
           IF #stringBox[#i] = #lineBreak THEN
               #lineBox[#pLineBox] := "Trim"(#lineBox[#pLineBox]);
               #pLineBox := #pLineBox + 1;
               #lineBox[#pLineBox] := #lineBreak;
               #pLineBox := #pLineBox + 1;
           END_IF;


           IF #stringBox[#i] <> #lineBreak THEN

               IF #i = 0 THEN
                   #lengthTest := #stringBox[#i];
               END_IF;

               IF #i >= 1 THEN
                   #lengthTest := CONCAT_WSTRING(IN1 := #lineBox[#pLineBox],
                                                 IN2 := #space,
                                                 IN3 := #stringBox[#i]);
               END_IF;

               IF LEN(#lengthTest) <= #maxLength THEN
                   #lineBox[#pLineBox] := #lengthTest;
               END_IF;

               IF LEN(#lengthTest) > #maxLength THEN
                   #lineBox[#pLineBox] := "Trim"(#lineBox[#pLineBox]);
                   #lineBox[#pLineBox] := "Trim"(#lineBox[#pLineBox]);
                   #pLineBox := #pLineBox + 1;
                   #lineBox[#pLineBox] := #stringBox[#i];
               END_IF;
           END_IF;

       END_FOR;

       FOR #i := 0 TO 10 DO

           IF #lineBox[#i] = #space OR #lineBox[#i] = WString#'' THEN
               EXIT;
           END_IF;
           IF #i = 0 THEN
               #output := #lineBox[#i];
           END_IF;
           IF #i >= 1 THEN
               IF #lineBox[#i] = #lineBreak THEN
                   #output := #output;
               END_IF;
               IF #lineBox[#i] <> #lineBreak THEN
                   #output := CONCAT_WSTRING(IN1 := #output,
                                             IN2 := #lineBreak,
                                             IN3 := #lineBox[#i]);
               END_IF;
           END_IF;

       END_FOR;

       #output := "Trim"(#output);

   END_IF;

   #"Word Wrap" := #output;
END_FUNCTION

FUNCTION "Trim" : WString   // FC29, SCL
{ S7_Optimized_Access := 'TRUE' }
VERSION : 0.1
   VAR_INPUT
      wString : WString;
   END_VAR
   VAR_TEMP
      ret : WString;
   END_VAR
   VAR CONSTANT
      space : WString := WSTRING#' ';
   END_VAR
BEGIN
   #ret := #wString;
   IF LEFT(IN := #ret, L := 1) = #space THEN
       #ret := RIGHT(IN := #ret, L := LEN(#ret) - 1);
   END_IF;
   IF RIGHT(IN := #ret, L := 1) = #space THEN
       #ret := LEFT(IN := #ret, L := LEN(#ret) - 1);
   END_IF;
   #Trim := #ret;
END_FUNCTION

FUNCTION "Upper" : Void   // FC49, SCL
{ S7_Optimized_Access := 'TRUE' }
VERSION : 0.1
   VAR_IN_OUT
      "string" : Variant;
   END_VAR
   VAR_TEMP
      "type" : Bool;
      stringBox : String;
      status : Int;
      wStringBox : WString;
      charArr : Array[0..255] of Char;
      cntChar : UInt;
      pChar : Int;
   END_VAR
   VAR CONSTANT
      asciiLow : Char := 'a';
      asciiHigh : Char := 'z';
      asciiCaseOffset : Int := 32;
   END_VAR
BEGIN
   IF TypeOf(#string) = String THEN
       #status := MOVE_BLK_VARIANT(SRC := #string,
                                   COUNT := 1,
                                   SRC_INDEX := 0,
                                   DEST_INDEX := 0,
                                   DEST => #stringBox);
   ELSIF TypeOf(#string) = WString THEN
       #status := MOVE_BLK_VARIANT(SRC := #string,
                                   COUNT := 1,
                                   SRC_INDEX := 0,
                                   DEST_INDEX := 0,
                                   DEST => #wStringBox);
       #stringBox := WSTRING_TO_STRING(#wStringBox);
   ELSE
       RETURN;
   END_IF;

   Strg_TO_Chars(Strg := #stringBox,
                 pChars := 0,
                 Cnt => #cntChar,
                 Chars := #charArr);

   FOR #pChar := 0 TO UINT_TO_INT(#cntChar) - 1 DO
       IF #asciiLow <= #charArr[#pChar] AND #charArr[#pChar] <= #asciiHigh THEN
           #charArr[#pChar] := INT_TO_CHAR(CHAR_TO_INT(#charArr[#pChar]) - #asciiCaseOffset);
       END_IF;
   END_FOR;

   Chars_TO_Strg(Chars := #charArr,
                 pChars := 0,
                 Cnt := #cntChar,
                 Strg => #stringBox);

   IF TypeOf(#string) = String THEN
       #status := MOVE_BLK_VARIANT(SRC := #stringBox,
                                   COUNT := 1,
                                   SRC_INDEX := 0,
                                   DEST_INDEX := 0,
                                   DEST => #string);
   ELSIF TypeOf(#string) = WString THEN
       #wStringBox := STRING_TO_WSTRING(#stringBox);
       #status := MOVE_BLK_VARIANT(SRC := #wStringBox,
                                   COUNT := 1,
                                   SRC_INDEX := 0,
                                   DEST_INDEX := 0,
                                   DEST => #string);
   END_IF;
END_FUNCTION

// folder: Utilities/Table Navigation

FUNCTION_BLOCK "Table Nav"   // FB43, SCL
{ S7_Optimized_Access := 'TRUE' }
VERSION : 0.1
   VAR_INPUT
      tblData : Variant;
      tblDisp : Variant;
      tableNav : "Table Nav: HMI";
   END_VAR
   VAR_IN_OUT
      rowIndices : Variant;
   END_VAR
   VAR
      "inst Pulses: Table Nav" : "Table Nav: Pulses";
      r1 : DInt;
   END_VAR
   VAR_TEMP
      len : Struct
         tblData : DInt;
         tblDisp : DInt;
      END_STRUCT;
      offset : DInt;
      pulses : "Table Nav: PLC";
      RET_VAL : Int;
      retRowIndices : Array[0..#lenRetArr] of DInt;
   END_VAR
   VAR CONSTANT
      lenRetArr : DInt := 999;
   END_VAR
BEGIN
   REGION "DESCRIPTION"
       (*
       The function returns row indicies indicating the visible rows of a larger
       table determined by standard table navigation buttons.
       The function uses the variant data type to handle tables of any size.
       Rollover and rollunder features are built in.
       *)    
   END_REGION

   REGION "GET PRESS PULSES"    
       #"inst Pulses: Table Nav"(press := #tableNav,
                                 pulses=> #pulses);
   END_REGION

   REGION "RUN ON BUTTON PRESS"
       IF "Table Nav: Run Trigger"(#pulses) THEN

           REGION "GET ARRAY PARAMETERS"
               #len.tblData := UDINT_TO_DINT(CountOfElements(#tblData));
               #len.tblDisp := UDINT_TO_DINT(CountOfElements(#tblDisp));
           END_REGION

           REGION "CALCULATE OFFSET"
               #offset := "Table Nav: Calculate Offset"(pulses := #pulses,
                                                        lenTblData := #len.tblData,
                                                        lenTblDisp := #len.tblDisp,
                                                        r1 := #r1);
           END_REGION

           REGION "CALCULATE FIRST ROW"
               #r1 := "Table Nav: Get First Row"(lenTblData := #len.tblData,
                                                 offset := #offset,
                                                 r1 := #r1);
           END_REGION

           REGION "CALCUALTE ROW INDICIES"
               "Table Nav: Calc Row Indices"(lenTblData := #len.tblData,
                                             lenTblDisp := #len.tblDisp,
                                             r1 := #r1,
                                             rowIndicies := #retRowIndices);
           END_REGION

           REGION "RETURN ROW INDICIES"
               #RET_VAL := MOVE_BLK_VARIANT(SRC := #retRowIndices,
                                            COUNT := DINT_TO_UDINT(#len.tblDisp),
                                            SRC_INDEX := 0,
                                            DEST_INDEX := 0,
                                            DEST => #rowIndices);
           END_REGION

       END_IF;
   END_REGION
END_FUNCTION_BLOCK

FUNCTION_BLOCK "Table Nav: Pulses"   // FB44, SCL
{ S7_Optimized_Access := 'TRUE' }
VERSION : 0.1
   VAR_INPUT
      press : "Table Nav: HMI";
   END_VAR
   VAR_OUTPUT
      pulses : "Table Nav: PLC";
   END_VAR
   VAR
      old : "Table Nav: PLC";
   END_VAR
BEGIN
   REGION "EVALUATION"
       #pulses.top := #press.top.actuate AND NOT #old.top;
       #pulses.pageUp := #press.pageUp.actuate AND NOT #old.pageUp;
       #pulses.lineUp := #press.lineUp.actuate AND NOT #old.lineUp;
       #pulses.lineDown := #press.lineDown.actuate AND NOT #old.lineDown;
       #pulses.pageDown := #press.pageDown.actuate AND NOT #old.pageDown;
       #pulses.bottom := #press.bottom.actuate AND NOT #old.bottom;
   END_REGION

   REGION "CHANGE DETECTION"
       #old.top := #press.top.actuate;
       #old.pageUp := #press.pageUp.actuate;
       #old.lineUp := #press.lineUp.actuate;
       #old.lineDown := #press.lineDown.actuate;
       #old.pageDown := #press.pageDown.actuate;
       #old.bottom := #press.bottom.actuate;
   END_REGION
END_FUNCTION_BLOCK

FUNCTION "Table Nav: Get First Row" : DInt   // FC44, SCL
{ S7_Optimized_Access := 'TRUE' }
VERSION : 0.1
   VAR_INPUT
      lenTblData : DInt;
      offset : DInt;
      r1 : DInt;
   END_VAR
   VAR_TEMP
      newR1 : DInt;
      trgRun : Bool;
   END_VAR
BEGIN
   REGION "DESCRIPTION"
       (*
       The new first row of the table is calculated from the offset. 
       Rollover and rollunder are resolved for the first row.
       *)
   END_REGION

   REGION "COPY TO INTERNAL"
       #newR1 := #r1 + #offset;
   END_REGION

   REGION "ROLLUNDER"
       IF #newR1 < 0 THEN
           #newR1 := #newR1 + #lenTblData;
       END_IF;
   END_REGION

   REGION "ROLLOVER"
       IF #newR1 > #lenTblData THEN
           #newR1 := #newR1 - #lenTblData;
       END_IF;
   END_REGION

   REGION "OUTPUT"
       #"Table Nav: Get First Row" := #newR1;
   END_REGION
END_FUNCTION

FUNCTION "Table Nav: Calculate Offset" : DInt   // FC45, SCL
{ S7_Optimized_Access := 'TRUE' }
VERSION : 0.1
   VAR_INPUT
      lenTblData : DInt;
      lenTblDisp : DInt;
      pulses : "Table Nav: PLC";
      r1 : DInt;
   END_VAR
   VAR_TEMP
      retOffset : DInt;
   END_VAR
   // Ret_Val : offset from table row 1 from button
BEGIN
   REGION "DESCRIPTION"
       (*
       The offset from the first row of the table is calculated based on the button pressed.
       *)
   END_REGION

   REGION "TOP"
       IF #pulses.top THEN
           #retOffset := -1 * #r1;
       END_IF;
   END_REGION

   REGION "PAGE UP"
       IF #pulses.pageUp THEN
           #retOffset := -1 * #lenTblDisp;
       END_IF;
   END_REGION

   REGION "LINE UP"
       IF #pulses.lineUp THEN
           #retOffset := -1;
       END_IF;
   END_REGION

   REGION "LINE DOWN"
       IF #pulses.lineDown THEN
           #retOffset := 1;
       END_IF;
   END_REGION

   REGION "PAGE DOWN"
       IF #pulses.pageDown THEN
           #retOffset := #lenTblDisp ;
       END_IF;
   END_REGION

   REGION "BOTTOM"
       IF #pulses.bottom THEN
           #retOffset := #lenTblData - #lenTblDisp - #r1;
       END_IF;
   END_REGION

   REGION "RETURN"
       #"Table Nav: Calculate Offset" := #retOffset;
   END_REGION
END_FUNCTION

FUNCTION "Table Nav: Calc Row Indices" : Void   // FC46, SCL
{ S7_Optimized_Access := 'TRUE' }
VERSION : 0.1
   VAR_INPUT
      lenTblData : DInt;
      lenTblDisp : DInt;
      r1 : DInt;
   END_VAR
   VAR_IN_OUT
      rowIndicies : Array[0..#lenRetArr] of DInt;
   END_VAR
   VAR_TEMP
      pOutArr : Int;
      calcRowIdx : DInt;
      retRowIndicies : Array[0..#lenRetArr] of DInt;
   END_VAR
   VAR CONSTANT
      lenRetArr : DInt := 999;
   END_VAR
BEGIN
   REGION "DESCRIPTION"
       (*
       An array of the row indicies that the table should display is returned.
       Rollover and rollunder are calculated index by index.
       *) 
   END_REGION

   REGION "INITIALIZE OUTPUT"
       FOR #pOutArr := 0 TO #lenRetArr DO
           #rowIndicies[#pOutArr] := 0;
       END_FOR;
   END_REGION

   REGION "CALCULATE INDICIES"
       FOR #pOutArr := 0 TO #lenTblDisp DO

           REGION "CALCULATE INDEX"
               #calcRowIdx := #r1 + #pOutArr;
           END_REGION

           REGION "ROLL UNDER"
               IF #calcRowIdx < 0 THEN
                   #calcRowIdx := #calcRowIdx + #lenTblDisp;
               END_IF;
           END_REGION

           REGION "ROLL OVER"
               IF #calcRowIdx >= #lenTblData THEN
                   #calcRowIdx := #calcRowIdx - #lenTblData;
               END_IF;
           END_REGION

           REGION "SAVE TO ARRAY"
               #retRowIndicies[#pOutArr] := #calcRowIdx;
           END_REGION

       END_FOR;
   END_REGION

   REGION "OUTPUT"
       #rowIndicies := #retRowIndicies;
   END_REGION
END_FUNCTION

FUNCTION "Table Nav: Run Trigger" : Bool   // FC47, SCL
{ S7_Optimized_Access := 'TRUE' }
VERSION : 0.1
   VAR_INPUT
      pulses : "Table Nav: PLC";
   END_VAR
BEGIN
       #"Table Nav: Run Trigger" :=
       #pulses.top OR
       #pulses.pageUp OR
       #pulses.lineUp OR
       #pulses.lineDown OR
       #pulses.pageDown OR
       #pulses.bottom;
END_FUNCTION

// folder: Utilities/Timer

FUNCTION "Timer: Time to WString" : WString   // FC36, SCL
{ S7_Optimized_Access := 'TRUE' }
VERSION : 0.1
   VAR_INPUT
      "Time" : Time;
   END_VAR
   VAR_TEMP
      "Time as DInt" : DInt;
      "Hours 10s Place" : DInt;
      "Hours 1s Place" : DInt;
      "Minutes 10s Place" : DInt;
      "Minutes 1s Place" : DInt;
      "Seconds 10s Place" : DInt;
      "Seconds 1s Place" : DInt;
      "Time Elements" : Array[0..4] of WString;
      Length : Int;
      "String Box" : WString;
      "DInt Box" : DInt;
   END_VAR
   VAR CONSTANT
      "Milliseconds per 10 Hours" : DInt := 36_000_000;
      "Milliseconds per Hour" : DInt := 3_600_000;
      "Milliseconds per 10 Minutes" : DInt := 600_000;
      "Milliseconds per Minute" : DInt := 60_000;
      "Milliseconds per 10 Seconds" : DInt := 10_000;
      "Milliseconds per Second" : DInt := 1_000;
   END_VAR
BEGIN
   REGION GET INPUT
       #"Time as DInt" := #Time;
   END_REGION

   REGION CONVERT TIME INTO INDIVIDUAL PLACE VALUES
       #"Minutes 10s Place" := #"Time as DInt" / #"Milliseconds per 10 Minutes";
       #"Minutes 1s Place" := (#"Time as DInt" / #"Milliseconds per Minute") MOD 10;
       #"Seconds 10s Place" := (#"Time as DInt" MOD #"Milliseconds per Minute") / #"Milliseconds per 10 Seconds";
       #"Seconds 1s Place" := (#"Time as DInt" / #"Milliseconds per Second") MOD 10;
   END_REGION

   REGION "ADD SIGN"
       #"Time Elements"[0] := wstring#'';
       IF #"Minutes 10s Place" < 0 OR
           #"Minutes 1s Place" < 0 OR
           #"Seconds 10s Place" < 0 OR
           #"Seconds 1s Place" < 0 THEN
            #"Time Elements"[0] := wstring#'-';
       END_IF;
   END_REGION

   REGION CONVERT PLACE VALUES INTO COMPONENT STRINGS
       // MINUTES
       #"DInt Box" := #"Minutes 10s Place" * 10 + #"Minutes 1s Place";
       #"String Box" := DINT_TO_WSTRING(IN := #"DInt Box");
       #"String Box" := "Strip Sign"("WString":=#"String Box");
       #"String Box" := "Add Leading"("Leading Character" := WCHAR#'0',
                                      "Desired Length" := 2,
                                      "String" := #"String Box");
       #"Time Elements"[1] := #"String Box";
       // COLON
       #"Time Elements"[2] := WSTRING#':';
       // SECONDS
       #"DInt Box" := #"Seconds 10s Place" * 10 + #"Seconds 1s Place";
       #"String Box" := DINT_TO_WSTRING(IN := #"DInt Box");
       #"String Box" := "Strip Sign"("WString":=#"String Box");
       #"String Box" := "Add Leading"("Leading Character" := WCHAR#'0',
                                      "Desired Length" := 2,
                                      "String" := #"String Box");
       #"Time Elements"[3] := #"String Box";
   END_REGION


   REGION RETURN VALUE
       #"Timer: Time to WString" := CONCAT_WSTRING(IN1 := #"Time Elements"[0],
                                            IN2 := #"Time Elements"[1],
                                            IN3 := #"Time Elements"[2],
                                            IN4 := #"Time Elements"[3]);
   END_REGION
END_FUNCTION

FUNCTION "Timer: WString to Time" : Time   // FC38, SCL
{ S7_Optimized_Access := 'TRUE' }
VERSION : 0.1
   VAR_INPUT
      WString : WString;
   END_VAR
   VAR_TEMP
      Count : UInt;
      "DInt Box" : DInt;
      "String Box" : WString [5];
      "Time Box" : Time;
      "WChar Array" : Array[0..4] of WChar;
   END_VAR
   VAR CONSTANT
      "ms/(10 hr)" : DInt := 36_000_000;
      "ms/hr" : DInt := 3_600_000;
      "ms/(10 min)" : DInt := 600_000;
      "ms/min" : DInt := 60_000;
      "ms/(10 sec)" : DInt := 10_000;
      "ms/sec" : DInt := 1_000;
   END_VAR
BEGIN
   REGION EXPLODE INPUT

       #"String Box" := #WString;
       IF #"String Box" = WSTRING#'' THEN
           #"String Box" := WSTRING#'00:00';
       END_IF;

       Strg_TO_Chars(Strg := #"String Box",
                     pChars := 0,
                     Cnt => #Count,
                     Chars := #"WChar Array");

   END_REGION

   REGION CONVERT ARRAY ELEMENTS TO TIME

       // 10S OF MINUTES
       #"DInt Box" := WCHAR_TO_DINT(IN := #"WChar Array"[0]) - 16#30;
       #"Time Box" := #"Time Box" + #"DInt Box" * #"ms/(10 min)";

       // MINUTES
       #"DInt Box" := WCHAR_TO_DINT(IN := #"WChar Array"[1]) - 16#30;
       #"Time Box" := #"Time Box" + #"DInt Box" * #"ms/min";

       // 10S OF SECONDS
       #"DInt Box" := WCHAR_TO_DINT(IN := #"WChar Array"[3]) - 16#30;
       #"Time Box" := #"Time Box" + #"DInt Box" * #"ms/(10 sec)";

       // SECONDS
       #"DInt Box" := WCHAR_TO_DINT(IN := #"WChar Array"[4]) - 16#30;
       #"Time Box" := #"Time Box" + #"DInt Box" * #"ms/sec";

   END_REGION


   REGION RETURN VALUE

       #"Timer: WString to Time" := #"Time Box";

   END_REGION
END_FUNCTION

FUNCTION "Timer: WString to Real" : Real   // FC39, SCL
{ S7_Optimized_Access := 'TRUE' }
VERSION : 0.1
   VAR_INPUT
      wstring : WString;
   END_VAR
   VAR CONSTANT
      msPerSec : Real := 1000.0;
   END_VAR
BEGIN
   #"Timer: WString to Real" := DINT_TO_REAL(TIME_TO_DINT("Timer: WString to Time"(#wstring))) / #msPerSec;
END_FUNCTION

FUNCTION "Timer: Real to WString" : WString   // FC40, SCL
{ S7_Optimized_Access := 'TRUE' }
VERSION : 0.1
   VAR_INPUT
      realVal : Real;
   END_VAR
   VAR CONSTANT
      msPerSec : Real := 1000.0;
   END_VAR
BEGIN
   #"Timer: Real to WString" := "Timer: Time to WString"(DINT_TO_TIME(REAL_TO_DINT(#realVal * #msPerSec)));
END_FUNCTION

// ===== library types =====

TYPE "Table Row Data"
   STRUCT
      address : UInt;
      ordered : Bool;
      pbSelection : Struct
         actuate : Bool;
         animate : USInt;
      END_STRUCT;
      rtBackground : Struct
         animate : USInt;
      END_STRUCT;
      tfDropZone : Struct
         animate : USInt;
         value : WString[20];
      END_STRUCT;
      tfLine : Struct
         animate : USInt;
         value : WString[20];
      END_STRUCT;
      tfPartNumber : Struct
         animateDL : USInt;
         animateSL : USInt;
         value : WString[40];
      END_STRUCT;
      tfTime : Struct
         animate : USInt;
         value : WString[20];
      END_STRUCT;
   END_STRUCT;
END_TYPE

TYPE "Station Assignment: Button Details Data"
   STRUCT
      alloted : Struct
         animate : USInt;
         value : WString[10];
      END_STRUCT;
      critical : Struct
         animate : USInt;
         value : WString[10];
      END_STRUCT;
      label : Struct
         animate : USInt;
         value : WString[2];
      END_STRUCT;
      partNumber : Struct
         animate : USInt;
         value : WString[40];
      END_STRUCT;
      select : Struct
         actuate : Bool;
         animate : USInt;
      END_STRUCT;
   END_STRUCT;
END_TYPE

TYPE "Station Sim Data"
   STRUCT
      stn : Struct
         animate : USInt;
         label : WString[20];
      END_STRUCT;
      btn : Struct
         actuate : Byte;
         animate : Array[0..7] of USInt;
         labels : Array[0..7] of WString [4];
      END_STRUCT;
   END_STRUCT;
END_TYPE

(* ===== HMI "HMI_RT_1" =====
system functions are stored by id; their names below are inferred from use
connection "Main HMI": ETHERNET, S7_1500_OMS

HMI tags "Default tag table"
   "Clock_Byte" : Byte = PLC Clock_Byte AT %MB0, 100 ms
   "HMI_screenNumber" : Int = PLC HMI.screenNumber AT %DB1.DBW0, 100 ms
   "HMI_barcode" : Barcode Screen = PLC HMI.barcode AT %DB1.DBW0, 100 ms
   "HMI_partCall_row{0}" : Table Row = PLC HMI.partCall.row[0], 100 ms
   "HMI_partCall_row{1}" : Table Row = PLC HMI.partCall.row[1], 100 ms
   "HMI_partCall_row{2}" : Table Row = PLC HMI.partCall.row[2], 100 ms
   "HMI_partCall_row{3}" : Table Row = PLC HMI.partCall.row[3], 100 ms
   "HMI_partCall_row{4}" : Table Row = PLC HMI.partCall.row[4], 100 ms
   "HMI_partCall_row{5}" : Table Row = PLC HMI.partCall.row[5], 100 ms
   "HMI_partCall_row{6}" : Table Row = PLC HMI.partCall.row[6], 100 ms
   "HMI_partCall_row{7}" : Table Row = PLC HMI.partCall.row[7], 100 ms
   "HMI_partCall_row{8}" : Table Row = PLC HMI.partCall.row[8], 100 ms
   "HMI_partCall_row{9}" : Table Row = PLC HMI.partCall.row[9], 100 ms
   "HMI_partCall_row{10}" : Table Row = PLC HMI.partCall.row[10], 100 ms
   "HMI_settings_stations_selectBtns{0}" : PB Data: Text Label = PLC HMI.settings.stations.selectBtns[0], 100 ms
   "HMI_settings_stations_selectBtns{1}" : PB Data: Text Label = PLC HMI.settings.stations.selectBtns[1], 100 ms
   "HMI_settings_stations_selectBtns{2}" : PB Data: Text Label = PLC HMI.settings.stations.selectBtns[2], 100 ms
   "HMI_settings_stations_selectBtns{3}" : PB Data: Text Label = PLC HMI.settings.stations.selectBtns[3], 100 ms
   "HMI_settings_stations_selectBtns{4}" : PB Data: Text Label = PLC HMI.settings.stations.selectBtns[4], 100 ms
   "HMI_settings_stations_selectBtns{5}" : PB Data: Text Label = PLC HMI.settings.stations.selectBtns[5], 100 ms
   "HMI_settings_stations_selectBtns{6}" : PB Data: Text Label = PLC HMI.settings.stations.selectBtns[6], 100 ms
   "HMI_settings_stations_selectBtns{7}" : PB Data: Text Label = PLC HMI.settings.stations.selectBtns[7], 100 ms
   "HMI_settings_stations_selectBtns{8}" : PB Data: Text Label = PLC HMI.settings.stations.selectBtns[8], 100 ms
   "HMI_settings_stations_selectBtns{9}" : PB Data: Text Label = PLC HMI.settings.stations.selectBtns[9], 100 ms
   "HMI_settings_stations_selectBtns{10}" : PB Data: Text Label = PLC HMI.settings.stations.selectBtns[10], 100 ms
   "HMI_settings_stations_selectBtns{11}" : PB Data: Text Label = PLC HMI.settings.stations.selectBtns[11], 100 ms
   "HMI_settings_kp8_buttons{0}" : PB Data: Text Label = PLC HMI.settings.kp8.buttons[0], 100 ms
   "HMI_settings_kp8_buttons{7}" : PB Data: Text Label = PLC HMI.settings.kp8.buttons[7], 100 ms
   "HMI_settings_kp8_buttons{3}" : PB Data: Text Label = PLC HMI.settings.kp8.buttons[3], 100 ms
   "HMI_settings_kp8_buttons{6}" : PB Data: Text Label = PLC HMI.settings.kp8.buttons[6], 100 ms
   "HMI_settings_kp8_buttons{2}" : PB Data: Text Label = PLC HMI.settings.kp8.buttons[2], 100 ms
   "HMI_settings_kp8_buttons{5}" : PB Data: Text Label = PLC HMI.settings.kp8.buttons[5], 100 ms
   "HMI_settings_kp8_buttons{1}" : PB Data: Text Label = PLC HMI.settings.kp8.buttons[1], 100 ms
   "HMI_settings_kp8_buttons{4}" : PB Data: Text Label = PLC HMI.settings.kp8.buttons[4], 100 ms
   "HMI_settings_stations_selCount" : Int = PLC HMI.settings.stations.selCount, 100 ms
   "HMI_settings_viewingStation_btns{0}" : Station: Assignment: Button Details = PLC HMI.settings.viewingStation.btns[0], 100 ms
   "HMI_settings_viewingStation_btns{1}" : Station: Assignment: Button Details = PLC HMI.settings.viewingStation.btns[1], 100 ms
   "HMI_settings_viewingStation_btns{2}" : Station: Assignment: Button Details = PLC HMI.settings.viewingStation.btns[2], 100 ms
   "HMI_settings_viewingStation_btns{3}" : Station: Assignment: Button Details = PLC HMI.settings.viewingStation.btns[3], 100 ms
   "HMI_settings_viewingStation_btns{4}" : Station: Assignment: Button Details = PLC HMI.settings.viewingStation.btns[4], 100 ms
   "HMI_settings_viewingStation_btns{5}" : Station: Assignment: Button Details = PLC HMI.settings.viewingStation.btns[5], 100 ms
   "HMI_settings_viewingStation_previous" : PB Data: Graphic/Text List = PLC HMI.settings.viewingStation.previous, 100 ms
   "HMI_settings_viewingStation_next" : PB Data: Graphic/Text List = PLC HMI.settings.viewingStation.next, 100 ms
   "HMI_settings_stations_selectAll" : PB Data: Text Label = PLC HMI.settings.stations.selectAll, 100 ms
   "HMI_settings_partNumber_assign" : PB Data: Text Label = PLC HMI.settings.partNumber.assign, 100 ms
   "HMI_settings_partNumber_ioField" : IO Field Data: Part Number = PLC HMI.settings.partNumber.ioField, 100 ms
   "HMI_settings_alotted_assign" : PB Data: Text Label = PLC HMI.settings.alotted.assign, 100 ms
   "HMI_settings_alotted_ioField" : IO Field Data: Timers = PLC HMI.settings.alotted.ioField, 100 ms
   "HMI_settings_critical_assign" : PB Data: Text Label = PLC HMI.settings.critical.assign, 100 ms
   "HMI_settings_critical_ioField" : IO Field Data: Timers = PLC HMI.settings.critical.ioField, 100 ms
   "HMI_settings_kp8_selectButtons" : PB Data: Text Label = PLC HMI.settings.kp8.selectButtons, 100 ms
   "HMI_settings_viewingStation_dzData" : Drop Zone Data = PLC HMI.settings.viewingStation.dzData, 100 ms
   "HMI_settings_viewingStation_lineData" : Line Label Data = PLC HMI.settings.viewingStation.lineData, 100 ms
   "HMI_settings_stations_prevGroup" : PB Data: Graphic/Text List = PLC HMI.settings.stations.prevGroup, 100 ms
   "HMI_settings_stations_nextGroup" : PB Data: Graphic/Text List = PLC HMI.settings.stations.nextGroup, 100 ms
   "HMI_settings_viewingStation_name" : WString[20] = PLC HMI.settings.viewingStation.name, 100 ms
   "HMI_tableNav_top" : PB Data: Graphic/Text List = PLC HMI.tableNav.top, 100 ms
   "HMI_tableNav_pageUp" : PB Data: Graphic/Text List = PLC HMI.tableNav.pageUp, 100 ms
   "HMI_tableNav_lineUp" : PB Data: Graphic/Text List = PLC HMI.tableNav.lineUp, 100 ms
   "HMI_tableNav_lineDown" : PB Data: Graphic/Text List = PLC HMI.tableNav.lineDown, 100 ms
   "HMI_tableNav_pageDown" : PB Data: Graphic/Text List = PLC HMI.tableNav.pageDown, 100 ms
   "HMI_tableNav_bottom" : PB Data: Graphic/Text List = PLC HMI.tableNav.bottom, 100 ms
   "HMI_simStations_stations{0}" : Station: Sim Data = PLC HMI.simStations.me[0] AT %DB1.DBX0.0, 100 ms
   "HMI_simStations_me{1}" : Station: Sim Data = PLC HMI.simStations.me[1], 100 ms
   "HMI_simStations_me{2}" : Station: Sim Data = PLC HMI.simStations.me[2], 100 ms
   "HMI_simStations_me{3}" : Station: Sim Data = PLC HMI.simStations.me[3], 100 ms
   "HMI_simStations_me{4}" : Station: Sim Data = PLC HMI.simStations.me[4], 100 ms
   "HMI_simStations_me{5}" : Station: Sim Data = PLC HMI.simStations.me[5], 100 ms
   "HMI_simStations_me{6}" : Station: Sim Data = PLC HMI.simStations.me[6], 100 ms
   "HMI_simStations_me{7}" : Station: Sim Data = PLC HMI.simStations.me[7], 100 ms
   "HMI_simStations_me{8}" : Station: Sim Data = PLC HMI.simStations.me[8], 100 ms
   "HMI_simStations_me{9}" : Station: Sim Data = PLC HMI.simStations.me[9], 100 ms
   "HMI_simStations_me{10}" : Station: Sim Data = PLC HMI.simStations.me[10], 100 ms
   "HMI_simStations_me{11}" : Station: Sim Data = PLC HMI.simStations.me[11], 100 ms
   "HMI_simStations_up" : PB Data: Graphic/Text List = PLC HMI.simStations.up, 100 ms
   "HMI_simStations_down" : PB Data: Graphic/Text List = PLC HMI.simStations.down, 100 ms
   "HMI_networkHealth_pnioDevices{1}" : PB Data: Text Label = PLC HMI.networkHealth.pnioDevices[1], 100 ms
   "HMI_networkHealth_pnioDevices{2}" : PB Data: Text Label = PLC HMI.networkHealth.pnioDevices[2], 100 ms
   "HMI_networkHealth_pnioDevices{3}" : PB Data: Text Label = PLC HMI.networkHealth.pnioDevices[3], 100 ms
   "HMI_networkHealth_pnioDevices{4}" : PB Data: Text Label = PLC HMI.networkHealth.pnioDevices[4], 100 ms
   "HMI_networkHealth_pnioDevices{5}" : PB Data: Text Label = PLC HMI.networkHealth.pnioDevices[5], 100 ms
   "HMI_networkHealth_pnioDevices{6}" : PB Data: Text Label = PLC HMI.networkHealth.pnioDevices[6], 100 ms
   "HMI_networkHealth_pnioDevices{7}" : PB Data: Text Label = PLC HMI.networkHealth.pnioDevices[7], 100 ms
   "HMI_networkHealth_pnioDevices{8}" : PB Data: Text Label = PLC HMI.networkHealth.pnioDevices[8], 100 ms
   "HMI_networkHealth_pnioDevices{9}" : PB Data: Text Label = PLC HMI.networkHealth.pnioDevices[9], 100 ms
   "HMI_networkHealth_pnioDevices{10}" : PB Data: Text Label = PLC HMI.networkHealth.pnioDevices[10], 100 ms
   "HMI_networkHealth_pnioDevices{11}" : PB Data: Text Label = PLC HMI.networkHealth.pnioDevices[11], 100 ms
   "HMI_networkHealth_pnioDevices{12}" : PB Data: Text Label = PLC HMI.networkHealth.pnioDevices[12], 100 ms
   "HMI_networkHealth_pnioDevices{13}" : PB Data: Text Label = PLC HMI.networkHealth.pnioDevices[13], 100 ms
   "HMI_networkHealth_pnioDevices{16}" : PB Data: Text Label = PLC HMI.networkHealth.pnioDevices[16], 100 ms
   "HMI_networkHealth_pnioDevices{14}" : PB Data: Text Label = PLC HMI.networkHealth.pnioDevices[14], 100 ms
   "HMI_networkHealth_pnioDevices{15}" : PB Data: Text Label = PLC HMI.networkHealth.pnioDevices[15], 100 ms
   "HMI_networkHealth_pnioDevices{17}" : PB Data: Text Label = PLC HMI.networkHealth.pnioDevices[17], 100 ms
   "HMI_networkHealth_pnioDevices{18}" : PB Data: Text Label = PLC HMI.networkHealth.pnioDevices[18], 100 ms
   "HMI_networkHealth_pnioDevices{19}" : PB Data: Text Label = PLC HMI.networkHealth.pnioDevices[19], 100 ms
   "HMI_networkHealth_pnioDevices{20}" : PB Data: Text Label = PLC HMI.networkHealth.pnioDevices[20], 100 ms
   "HMI_networkHealth_pnioDevices{21}" : PB Data: Text Label = PLC HMI.networkHealth.pnioDevices[21], 100 ms
   "HMI_networkHealth_pnioDevices{22}" : PB Data: Text Label = PLC HMI.networkHealth.pnioDevices[22], 100 ms
   "HMI_networkHealth_pnioDevices{31}" : PB Data: Text Label = PLC HMI.networkHealth.pnioDevices[31], 100 ms
   "HMI_networkHealth_pnioDevices{32}" : PB Data: Text Label = PLC HMI.networkHealth.pnioDevices[32], 100 ms
   "HMI_networkHealth_pnioDevices{29}" : PB Data: Text Label = PLC HMI.networkHealth.pnioDevices[29], 100 ms
   "HMI_networkHealth_pnioDevices{30}" : PB Data: Text Label = PLC HMI.networkHealth.pnioDevices[30], 100 ms
   "HMI_networkHealth_pnioDevices{27}" : PB Data: Text Label = PLC HMI.networkHealth.pnioDevices[27], 100 ms
   "HMI_networkHealth_pnioDevices{28}" : PB Data: Text Label = PLC HMI.networkHealth.pnioDevices[28], 100 ms
   "HMI_networkHealth_pnioDevices{23}" : PB Data: Text Label = PLC HMI.networkHealth.pnioDevices[23], 100 ms
   "HMI_networkHealth_pnioDevices{24}" : PB Data: Text Label = PLC HMI.networkHealth.pnioDevices[24], 100 ms
   "HMI_networkHealth_pnioDevices{25}" : PB Data: Text Label = PLC HMI.networkHealth.pnioDevices[25], 100 ms
   "HMI_networkHealth_pnioDevices{26}" : PB Data: Text Label = PLC HMI.networkHealth.pnioDevices[26], 100 ms
   "HMI_networkHealth_pnioDevices{33}" : PB Data: Text Label = PLC HMI.networkHealth.pnioDevices[33], 100 ms
   "HMI_networkHealth_pnioDevices{34}" : PB Data: Text Label = PLC HMI.networkHealth.pnioDevices[34], 100 ms
   "HMI_networkHealth_pnioDevices{35}" : PB Data: Text Label = PLC HMI.networkHealth.pnioDevices[35], 100 ms
   "HMI_networkHealth_pnioDevices{36}" : PB Data: Text Label = PLC HMI.networkHealth.pnioDevices[36], 100 ms
   "HMI_networkHealth_pnioDevices{37}" : PB Data: Text Label = PLC HMI.networkHealth.pnioDevices[37], 100 ms
   "HMI_networkHealth_pnioDevices{38}" : PB Data: Text Label = PLC HMI.networkHealth.pnioDevices[38], 100 ms
   "HMI_networkHealth_pnioDevices{39}" : PB Data: Text Label = PLC HMI.networkHealth.pnioDevices[39], 100 ms
   "HMI_networkHealth_pnioDevices{40}" : PB Data: Text Label = PLC HMI.networkHealth.pnioDevices[40], 100 ms
   "HMI_networkHealth_pnioDevices{41}" : PB Data: Text Label = PLC HMI.networkHealth.pnioDevices[41], 100 ms
   "HMI_networkHealth_pnioDevices{42}" : PB Data: Text Label = PLC HMI.networkHealth.pnioDevices[42], 100 ms
   "HMI_networkHealth_pnioDevices{43}" : PB Data: Text Label = PLC HMI.networkHealth.pnioDevices[43], 100 ms
   "HMI_networkHealth_pnioDevices{44}" : PB Data: Text Label = PLC HMI.networkHealth.pnioDevices[44], 100 ms
   "HMI_networkHealth_pnioDevices{45}" : PB Data: Text Label = PLC HMI.networkHealth.pnioDevices[45], 100 ms
   "HMI_networkHealth_pnioDevices{46}" : PB Data: Text Label = PLC HMI.networkHealth.pnioDevices[46], 100 ms
   "HMI_networkHealth_pnioDevices{47}" : PB Data: Text Label = PLC HMI.networkHealth.pnioDevices[47], 100 ms
   "HMI_networkHealth_pnioDevices{48}" : PB Data: Text Label = PLC HMI.networkHealth.pnioDevices[48], 100 ms
   "HMI_networkHealth_et200spPopUp" : Station: ET200SP Comm Debug Data = PLC HMI.networkHealth.et200spPopUp, 100 ms
   "HMI_networkHealth_kp8PopUp" : Station: KP8 Comm Debug Data = PLC HMI.networkHealth.kp8PopUp, 100 ms
   "HMI_networkHealth_selectedDevice" : Int = PLC HMI.networkHealth.selectedDevice, 100 ms
   "Recipe Buffer_dropZone" : USInt = PLC "Recipe Buffer".dropZone, 1 s
   "Recipe Buffer_kp8Output" : DWord = PLC "Recipe Buffer".kp8Output, 1 s
   "Recipe Buffer_kp8LogicalState0" : Bool = PLC "Recipe Buffer".kp8LogicalState0, 1 s
   "Recipe Buffer_kp8LogicalState1" : Bool = PLC "Recipe Buffer".kp8LogicalState1, 1 s
   "Recipe Buffer_kp8LogicalState2" : Bool = PLC "Recipe Buffer".kp8LogicalState2, 1 s
   "Recipe Buffer_kp8LogicalState3" : Bool = PLC "Recipe Buffer".kp8LogicalState3, 1 s
   "Recipe Buffer_kp8LogicalState4" : Bool = PLC "Recipe Buffer".kp8LogicalState4, 1 s
   "Recipe Buffer_kp8LogicalState5" : Bool = PLC "Recipe Buffer".kp8LogicalState5, 1 s
   "Recipe Buffer_kp8LogicalState6" : Bool = PLC "Recipe Buffer".kp8LogicalState6, 1 s
   "Recipe Buffer_kp8LogicalState7" : Bool = PLC "Recipe Buffer".kp8LogicalState7, 1 s
   "Recipe Buffer_lineName" : USInt = PLC "Recipe Buffer".lineName, 1 s
   "Recipe Buffer_pnCode" : DInt = PLC "Recipe Buffer".pnCode, 1 s
   "Recipe Buffer_stackLight" : DWord = PLC "Recipe Buffer".stackLight, 1 s
   "Recipe Buffer_wipName" : WString[254] = PLC "Recipe Buffer".wipName, 1 s
   "Recipe Buffer_wipNumber" : UInt = PLC "Recipe Buffer".wipNumber, 1 s

text list "Station Selection Single": 0 'Select a Station to View'; 1 'Assignments'

recipe "Station01": dz <- "Recipe Buffer_dropZone", kp8Output <- "Recipe Buffer_kp8Output", logicalState0 <- "Recipe Buffer_kp8LogicalState0", logicalState1 <- "Recipe Buffer_kp8LogicalState1", logicalState2 <- "Recipe Buffer_kp8LogicalState2", logicalState3 <- "Recipe Buffer_kp8LogicalState3", logicalState4 <- "Recipe Buffer_kp8LogicalState4", logicalState5 <- "Recipe Buffer_kp8LogicalState5", logicalState6 <- "Recipe Buffer_kp8LogicalState6", logicalState7 <- "Recipe Buffer_kp8LogicalState7", lineName <- "Recipe Buffer_lineName", pnCode <- "Recipe Buffer_pnCode", stackLight <- "Recipe Buffer_stackLight", wipName <- "Recipe Buffer_wipName", wipNumber <- "Recipe Buffer_wipNumber"

recipe "Station02": dz <- "Recipe Buffer_dropZone", kp8Output <- "Recipe Buffer_kp8Output", logicalState0 <- "Recipe Buffer_kp8LogicalState0", logicalState1 <- "Recipe Buffer_kp8LogicalState1", logicalState2 <- "Recipe Buffer_kp8LogicalState2", logicalState3 <- "Recipe Buffer_kp8LogicalState3", logicalState4 <- "Recipe Buffer_kp8LogicalState4", logicalState5 <- "Recipe Buffer_kp8LogicalState5", logicalState6 <- "Recipe Buffer_kp8LogicalState6", logicalState7 <- "Recipe Buffer_kp8LogicalState7", lineName <- "Recipe Buffer_lineName", pnCode <- "Recipe Buffer_pnCode", stackLight <- "Recipe Buffer_stackLight", wipName <- "Recipe Buffer_wipName", wipNumber <- "Recipe Buffer_wipNumber"

recipe "Station03": dz <- "Recipe Buffer_dropZone", kp8Output <- "Recipe Buffer_kp8Output", logicalState0 <- "Recipe Buffer_kp8LogicalState0", logicalState1 <- "Recipe Buffer_kp8LogicalState1", logicalState2 <- "Recipe Buffer_kp8LogicalState2", logicalState3 <- "Recipe Buffer_kp8LogicalState3", logicalState4 <- "Recipe Buffer_kp8LogicalState4", logicalState5 <- "Recipe Buffer_kp8LogicalState5", logicalState6 <- "Recipe Buffer_kp8LogicalState6", logicalState7 <- "Recipe Buffer_kp8LogicalState7", lineName <- "Recipe Buffer_lineName", pnCode <- "Recipe Buffer_pnCode", stackLight <- "Recipe Buffer_stackLight", wipName <- "Recipe Buffer_wipName", wipNumber <- "Recipe Buffer_wipNumber"

recipe "Station04": dz <- "Recipe Buffer_dropZone", kp8Output <- "Recipe Buffer_kp8Output", logicalState0 <- "Recipe Buffer_kp8LogicalState0", logicalState1 <- "Recipe Buffer_kp8LogicalState1", logicalState2 <- "Recipe Buffer_kp8LogicalState2", logicalState3 <- "Recipe Buffer_kp8LogicalState3", logicalState4 <- "Recipe Buffer_kp8LogicalState4", logicalState5 <- "Recipe Buffer_kp8LogicalState5", logicalState6 <- "Recipe Buffer_kp8LogicalState6", logicalState7 <- "Recipe Buffer_kp8LogicalState7", lineName <- "Recipe Buffer_lineName", pnCode <- "Recipe Buffer_pnCode", stackLight <- "Recipe Buffer_stackLight", wipName <- "Recipe Buffer_wipName", wipNumber <- "Recipe Buffer_wipNumber"

recipe "Station05": dz <- "Recipe Buffer_dropZone", kp8Output <- "Recipe Buffer_kp8Output", logicalState0 <- "Recipe Buffer_kp8LogicalState0", logicalState1 <- "Recipe Buffer_kp8LogicalState1", logicalState2 <- "Recipe Buffer_kp8LogicalState2", logicalState3 <- "Recipe Buffer_kp8LogicalState3", logicalState4 <- "Recipe Buffer_kp8LogicalState4", logicalState5 <- "Recipe Buffer_kp8LogicalState5", logicalState6 <- "Recipe Buffer_kp8LogicalState6", logicalState7 <- "Recipe Buffer_kp8LogicalState7", lineName <- "Recipe Buffer_lineName", pnCode <- "Recipe Buffer_pnCode", stackLight <- "Recipe Buffer_stackLight", wipName <- "Recipe Buffer_wipName", wipNumber <- "Recipe Buffer_wipNumber"

recipe "Station06": dz <- "Recipe Buffer_dropZone", kp8Output <- "Recipe Buffer_kp8Output", logicalState0 <- "Recipe Buffer_kp8LogicalState0", logicalState1 <- "Recipe Buffer_kp8LogicalState1", logicalState2 <- "Recipe Buffer_kp8LogicalState2", logicalState3 <- "Recipe Buffer_kp8LogicalState3", logicalState4 <- "Recipe Buffer_kp8LogicalState4", logicalState5 <- "Recipe Buffer_kp8LogicalState5", logicalState6 <- "Recipe Buffer_kp8LogicalState6", logicalState7 <- "Recipe Buffer_kp8LogicalState7", lineName <- "Recipe Buffer_lineName", pnCode <- "Recipe Buffer_pnCode", stackLight <- "Recipe Buffer_stackLight", wipName <- "Recipe Buffer_wipName", wipNumber <- "Recipe Buffer_wipNumber"

screen "1 PART CALL" 1366x768
   on GenerateScreen: SetTag("HMI_screenNumber", 1)
   Rectangle "Settings Tab Background" at 682,0 size 684x68
      Appearance <- "HMI_screenNumber"
   Rectangle "Part Call Tab Background" at 0,0 size 685x68
      Appearance <- "HMI_screenNumber"
   Rectangle "Settings Tab Border Hide" at 685,61 size 678x20
      Visibility <- "HMI_screenNumber"
   Rectangle "Part Call Tab Border Hide" at 3,61 size 679x20
      Visibility <- "HMI_screenNumber"
   Button "Settings Screen" at 683,0 size 683x68; TextOff 'SETTINGS'; Authorization "User administration"
      on Release: ActivateScreen("2 SETTINGS", 0)
   Button "Part Call Screen" at 0,0 size 683x68; TextOff 'PART CALL'
      on Release: ActivateScreen("1 PART CALL", 0)
   TextField "Header Line" at 32,112 size 216x53; Text 'LINE'
   TextField "Header Drop Zone" at 238,112 size 236x53; Text 'DROP ZONE'
   TextField "Header Part Number" at 474,112 size 648x53; Text 'PART NUMBER'
   TextField "Header Time" at 1112,112 size 222x53; Text 'TIME'
   ScreenModuleView "TableRow00" at 27,170 size 1312x52; ScreenModuleType ""
      Guid_{11997190-27688} <- "HMI_partCall_row{0}"
      on Guid_{11997190-83214}: ActivateScreen("3 BARCODE", 0)
   ScreenModuleView "TableRow01" at 27,222 size 1312x52; ScreenModuleType ""
      Guid_{11997190-27688} <- "HMI_partCall_row{1}"
      on Guid_{11997190-83214}: ActivateScreen("3 BARCODE", 0)
   ScreenModuleView "TableRow02" at 27,274 size 1312x52; ScreenModuleType ""
      Guid_{11997190-27688} <- "HMI_partCall_row{2}"
      on Guid_{11997190-83214}: ActivateScreen("3 BARCODE", 0)
   ScreenModuleView "TableRow03" at 27,326 size 1312x52; ScreenModuleType ""
      Guid_{11997190-27688} <- "HMI_partCall_row{3}"
      on Guid_{11997190-83214}: ActivateScreen("3 BARCODE", 0)
   ScreenModuleView "TableRow04" at 27,378 size 1312x52; ScreenModuleType ""
      Guid_{11997190-27688} <- "HMI_partCall_row{4}"
      on Guid_{11997190-83214}: ActivateScreen("3 BARCODE", 0)
   ScreenModuleView "TableRow05" at 27,430 size 1312x52; ScreenModuleType ""
      Guid_{11997190-27688} <- "HMI_partCall_row{5}"
      on Guid_{11997190-83214}: ActivateScreen("3 BARCODE", 0)
   ScreenModuleView "TableRow06" at 27,482 size 1312x52; ScreenModuleType ""
      Guid_{11997190-27688} <- "HMI_partCall_row{6}"
      on Guid_{11997190-83214}: ActivateScreen("3 BARCODE", 0)
   ScreenModuleView "TableRow07" at 27,534 size 1312x52; ScreenModuleType ""
      Guid_{11997190-27688} <- "HMI_partCall_row{7}"
      on Guid_{11997190-83214}: ActivateScreen("3 BARCODE", 0)
   ScreenModuleView "TableRow08" at 27,586 size 1312x52; ScreenModuleType ""
      Guid_{11997190-27688} <- "HMI_partCall_row{8}"
      on Guid_{11997190-83214}: ActivateScreen("3 BARCODE", 0)
   ScreenModuleView "TableRow09" at 27,638 size 1312x52; ScreenModuleType ""
      Guid_{11997190-27688} <- "HMI_partCall_row{9}"
      on Guid_{11997190-83214}: ActivateScreen("3 BARCODE", 0)
   ScreenModuleView "TableRow10" at 27,690 size 1312x52; ScreenModuleType ""
      Guid_{11997190-27688} <- "HMI_partCall_row{10}"
      on Guid_{11997190-83214}: ActivateScreen("3 BARCODE", 0)

screen "2 SETTINGS" 1366x768
   on GenerateScreen: SetTag("HMI_screenNumber", 2)
   Rectangle "Part Call Nave Panel" at 0,0 size 455x68
      Appearance <- "HMI_screenNumber"
   Rectangle "Settings Nav Panel" at 452,0 size 462x68
      Appearance <- "HMI_screenNumber"
   Rectangle "Network Health Nav Panel" at 911,0 size 455x68
      Appearance <- "HMI_screenNumber"
   Rectangle "Part Call Border Hide" at 3,60 size 449x20
      Visibility <- "HMI_screenNumber"
   Rectangle "Settings Border Hide" at 455,60 size 456x20
      Visibility <- "HMI_screenNumber"
   Rectangle "Network Health Border Hide" at 914,60 size 449x20
      Visibility <- "HMI_screenNumber"
   Button "Part Call Screen" at 0,0 size 455x68; TextOff 'PART CALL'
      on Release: ActivateScreen("1 PART CALL", 0)
   Button "Settings Screen" at 455,0 size 460x68; TextOff 'SETTINGS'
      on Release: ActivateScreen("2 SETTINGS", 0)
   Button "Network Health Screen" at 914,0 size 452x68; TextOff 'NW HEALTH'
      on Release: ActivateScreen("4 NETWORK HEALTH", 0)
   Rectangle "Station Assignment Table BG Full" at 793,120 size 533x630
      Visibility <- "HMI_settings_stations_selCount"
   TextField "Current Station Single" at 803,130 size 513x45; Text 'Text'
      Visibility <- "HMI_settings_stations_selCount"
   TextField "Hide Line and Drop Zone Multi" at 803,181 size 513x40; Text 'select single station for Line and Drop Zone'
      Visibility <- "HMI_settings_stations_selCount"
   GraphicView "KP8 Image" at 496,327 size 275x412; Picture "kp8 image"
   Rectangle "Station Assignment Table BG Mini" at 793,120 size 533x65
      Visibility <- "HMI_settings_stations_selCount"
   ScreenModuleView "PB: Set PN" at 50,130 size 414x45; Guid_{11997190-63616} 'Assign Part Number'; ScreenModuleType ""
      Guid_{11997190-63605} <- "HMI_settings_partNumber_assign"
   ScreenModuleView "PN IO Field" at 50,180 size 414x50; ScreenModuleType ""
      Guid_{11997190-63113} <- "HMI_settings_partNumber_ioField"
   ScreenModuleView "PB: Set Allotted" at 494,130 size 137x45; Guid_{11997190-63616} 'Allotted'; ScreenModuleType ""
      Guid_{11997190-63605} <- "HMI_settings_alotted_assign"
   ScreenModuleView "PB: Set Critical" at 636,130 size 137x45; Guid_{11997190-63616} 'Crititcal'; ScreenModuleType ""
      Guid_{11997190-63605} <- "HMI_settings_critical_assign"
   ScreenModuleView "Alotted Time IO Field" at 494,180 size 137x50; ScreenModuleType ""
      Guid_{11997190-63269} <- "HMI_settings_alotted_ioField"
   ScreenModuleView "Critical Time IO Field" at 636,180 size 137x50; ScreenModuleType ""
      Guid_{11997190-63269} <- "HMI_settings_critical_ioField"
   ScreenModuleView "PB: Select KP8 Buttons" at 493,270 size 284x45; Guid_{11997190-63616} 'Select Buttons'; ScreenModuleType ""
      Guid_{11997190-63605} <- "HMI_settings_kp8_selectButtons"
   ScreenModuleView "KP8 00: RESET" at 641,614 size 68x66; ScreenModuleType ""
      Guid_{11997190-57808} <- "HMI_settings_kp8_buttons{0}"
   ScreenModuleView "KP8 01" at 641,535 size 68x66; ScreenModuleType ""
      Guid_{11997190-57808} <- "HMI_settings_kp8_buttons{1}"
   ScreenModuleView "KP8 02" at 641,459 size 68x66; ScreenModuleType ""
      Guid_{11997190-57808} <- "HMI_settings_kp8_buttons{2}"
   ScreenModuleView "KP8 03" at 641,383 size 68x66; ScreenModuleType ""
      Guid_{11997190-57808} <- "HMI_settings_kp8_buttons{3}"
   ScreenModuleView "KP8 04: STOP RUNTIME" at 557,614 size 68x66; ScreenModuleType ""
      on Guid_{11997190-59171}: StopRuntime(0)
      Guid_{11997190-57808} <- "HMI_settings_kp8_buttons{4}"
   ScreenModuleView "KP8 05" at 557,535 size 68x66; ScreenModuleType ""
      Guid_{11997190-57808} <- "HMI_settings_kp8_buttons{5}"
   ScreenModuleView "KP8 06" at 557,459 size 68x66; ScreenModuleType ""
      Guid_{11997190-57808} <- "HMI_settings_kp8_buttons{6}"
   ScreenModuleView "KP8 07" at 557,383 size 68x66; ScreenModuleType ""
      Guid_{11997190-57808} <- "HMI_settings_kp8_buttons{7}"
   ScreenModuleView "PB: Previous Group" at 50,270 size 65x45; Guid_{11997190-63799} "Up"; ScreenModuleType ""
      Guid_{11997190-63779} <- "HMI_settings_stations_prevGroup"
   ScreenModuleView "PB: Select All Stations" at 120,270 size 274x45; Guid_{11997190-63616} 'Select Stations'; ScreenModuleType ""
      Guid_{11997190-63605} <- "HMI_settings_stations_selectAll"
   ScreenModuleView "PB: Next Group" at 399,270 size 65x45; Guid_{11997190-63799} "Down"; ScreenModuleType ""
      Guid_{11997190-63779} <- "HMI_settings_stations_nextGroup"
   ScreenModuleView "Station 00 Select" at 50,320 size 205x65; ScreenModuleType ""
      Guid_{11997190-57808} <- "HMI_settings_stations_selectBtns{0}"
   ScreenModuleView "Station 01 Select" at 260,320 size 205x65; ScreenModuleType ""
      Guid_{11997190-57808} <- "HMI_settings_stations_selectBtns{1}"
   ScreenModuleView "Station 02 Select" at 50,391 size 205x65; ScreenModuleType ""
      Guid_{11997190-57808} <- "HMI_settings_stations_selectBtns{2}"
   ScreenModuleView "Station 03 Select" at 260,391 size 205x65; ScreenModuleType ""
      Guid_{11997190-57808} <- "HMI_settings_stations_selectBtns{3}"
   ScreenModuleView "Station 04 Select" at 50,462 size 205x65; ScreenModuleType ""
      Guid_{11997190-57808} <- "HMI_settings_stations_selectBtns{4}"
   ScreenModuleView "Station 05 Select" at 260,462 size 205x65; ScreenModuleType ""
      Guid_{11997190-57808} <- "HMI_settings_stations_selectBtns{5}"
   ScreenModuleView "Station 06 Select" at 50,533 size 205x65; ScreenModuleType ""
      Guid_{11997190-57808} <- "HMI_settings_stations_selectBtns{6}"
   ScreenModuleView "Station 07 Select" at 260,533 size 205x65; ScreenModuleType ""
      Guid_{11997190-57808} <- "HMI_settings_stations_selectBtns{7}"
   ScreenModuleView "Station 08 Select" at 50,604 size 205x65; ScreenModuleType ""
      Guid_{11997190-57808} <- "HMI_settings_stations_selectBtns{8}"
   ScreenModuleView "Station 09 Select" at 260,604 size 205x65; ScreenModuleType ""
      Guid_{11997190-57808} <- "HMI_settings_stations_selectBtns{9}"
   ScreenModuleView "Station 10 Select" at 50,675 size 205x65; ScreenModuleType ""
      Guid_{11997190-57808} <- "HMI_settings_stations_selectBtns{10}"
   ScreenModuleView "Station 11 Select" at 260,675 size 205x65; ScreenModuleType ""
      Guid_{11997190-57808} <- "HMI_settings_stations_selectBtns{11}"
   ScreenModuleView "Line Label" at 803,181 size 267x40; ScreenModuleType ""
      Guid_{11997190-64598} <- "HMI_settings_viewingStation_lineData"
   ScreenModuleView "Drop Zone Label" at 1076,181 size 240x40; ScreenModuleType ""
      Guid_{11997190-64802} <- "HMI_settings_viewingStation_dzData"
   ScreenModuleView "PB: Previous Station" at 803,130 size 65x45; Guid_{11997190-63799} "Left"; ScreenModuleType ""
      Guid_{11997190-63779} <- "HMI_settings_viewingStation_previous"
   TextField "Current Station Multi" at 873,130 size 373x45; Text 'Assignments'
      Visibility <- "HMI_settings_stations_selCount"
   ScreenModuleView "PB: Next Station" at 1251,130 size 65x45; Guid_{11997190-63799} "Right"; ScreenModuleType ""
      Guid_{11997190-63779} <- "HMI_settings_viewingStation_next"
   TextField "Button Column Header" at 803,226 size 75x40; Text 'Btn'
      Visibility <- "HMI_settings_stations_selCount"
   TextField "Timer Column Header" at 872,226 size 128x40; Text 'Times'
      Visibility <- "HMI_settings_stations_selCount"
   TextField "Part Number Column Header" at 993,226 size 323x40; Text 'Part Number'
      Visibility <- "HMI_settings_stations_selCount"
   ScreenModuleView "Button 00 Details" at 803,271 size 513x74; ScreenModuleType ""
      Guid_{11997190-60358} <- "HMI_settings_viewingStation_btns{0}"
   ScreenModuleView "Button 01 Details" at 803,350 size 513x74; ScreenModuleType ""
      Guid_{11997190-60358} <- "HMI_settings_viewingStation_btns{1}"
   ScreenModuleView "Button 02 Details" at 803,429 size 513x74; ScreenModuleType ""
      Guid_{11997190-60358} <- "HMI_settings_viewingStation_btns{2}"
   ScreenModuleView "Button 03 Details" at 803,508 size 513x74; ScreenModuleType ""
      Guid_{11997190-60358} <- "HMI_settings_viewingStation_btns{3}"
   ScreenModuleView "Button 04 Details" at 803,587 size 513x74; ScreenModuleType ""
      Guid_{11997190-60358} <- "HMI_settings_viewingStation_btns{4}"
   ScreenModuleView "Button 05 Details" at 803,666 size 513x74; ScreenModuleType ""
      Guid_{11997190-60358} <- "HMI_settings_viewingStation_btns{5}"

